
text list "Disconnect Code Descriptions Long": 0 'Connection terminated successfully.'; 28672 'No job processing active.'; 28673 'Start of job processing, connection being terminated.'; 28674 'Intermediate call (REQ irrelevant), connection being terminated.'; 32902 'The ID parameter is not in the permitted value range.'; 32931 'Attempt is being made to terminate a non-existent connection or the connection is already terminated.'; 32964 'Temporary communication error: New parameters are being assigned to the interface or the connection is currently being established.'; 65535 'In connect state.'

text list "Send Code Descriptions Long": 0 'Send job completed without error.'; 28672 'No job processing active.'; 28673 'Start of job execution, data is being sent. When processing this job, the operating system accesses the data in the DATA send area.'; 28674 'Job executing (REQ irrelevant). When processing this job, the operating system accesses the data in the DATA send area.'; 32901 'The LEN parameter is greater than the highest permitted value (65536). DATA and LEN parameters both have the value "0".'; 32902 'The ID parameter is outside the permitted address range (1..0xFFF).'; 32904 'The LEN parameter is greater than the area specified in DATA.'; 32929 'Communication error: The specified connection has not yet been established. The specified connection is being terminated. Transfer via thisconnection is not possible. The interface is being re-initialized.'; 32947 'The protocol variant (ConnectionType parameter in the connection description) is set to UDP. Use the instruction "TUSEND" with a UDP connection.'; 32963 'A block with this ID is already being processed in a different priority group. Internal lack of resources.'; 32964 'Temporary communication error: The connection cannot be established to the partner at this time. The interface is receiving new parameter settings or the connection is being established.'; 32965 'Connection terminated by the communication partner.'; 32966 'Network error. Communication partner cannot be reached.'; 32967 'Execution timeout'; 65535 'Function not yet called.'

text list "Status Lists": 0 ''; 1 ''; 2 ''; 3 ''

ScreenModuleEditorView "Connection_Status_Details" 790x405
   SymbolicIOField "header" at 0,0 size 790x50; TextOn '1'; TextOff '0'; TextList "Connection Details Header"
      Appearance <- "interface.header_animate"
      Visibility <- "interface.header_visible"
      ProcessValue <- "interface.header_selector"
   IOField "payload" at 0,55 size 790x295; FormatPattern ?????????????????????????????????????????????????????????????????????????????????????????????????????????????????????????????????????????????????????????????????????????????????????????????????????????????????????????????????????????????????????????????
      ProcessValue <- "interface.payload_text"
      Appearance <- "interface.payload_animate"
      Visibility <- "interface.payload_visible"
   Button "display_payload_button" at 0,355 size 790x50; TextOff 'DISPLAY PAYLOAD'
      Appearance <- "interface.display_payload_button_animate"
      ObjectEnable <- "interface.display_payload_button_enable"
      Visibility <- "interface.display_payload_button_visible"
      on Press: function_b14e0dd5("interface.display_payload_button_actuate", 0)
   SymbolicIOField "detailed_status" at 0,55 size 790x295; TextOff '0'; TextOn '1'; TextList "Status Lists"
      ProcessValue <- "interface.detailed_status_list_selector"
      Visibility <- "interface.detailed_status_visible"
      Appearance <- "interface.detailed_status_animate"
   Button "back_button" at 0,0 size 790x405; TextOff 'Text'
      ObjectEnable <- "interface.back_button_enable"
      Visibility <- "interface.back_button_visible"
      on Press: function_b14e0dd5("interface.back_button_actuate", 0)
*)

(* ===== HMI "HMI_RT_1" =====
system functions are stored by id; their names below are inferred from use

text list "Connection Details Header": 0 'NO STATE'; 1 'DISCONNECTION STATUS'; 2 'CONNECTION STATUS'; 3 'SEND STATUS'

text list "Connect Code Descriptions Long": 0 'Connection successfully established.'; 28672 'No job processing active'; 28673 'Start job execution, establish connection.'; 28674 'Connection is being established (REQ irrelevant).'; 32901 'Connection ID (ID parameter) is already being used by a configured connection.'; 32902 'The ID parameter is outside the valid range.'; 32903 'Maximum number of connections reached; no additional connection possible'; 32905 'The CONNECT parameter does not point to a data block.'; 32922 'The structure at the CONNECT parameter is not supported on an integrated interface or the length is invalid or an incorrect "InterfaceID" is specified in the connection description (SDT).'; 32923 'The element InterfaceId within the TCON_xxx structure does not reference a hardware identifier of a CPU or CM/CP interface or has the value "0".'; 32928 'Group error for error codes W#16#80A1 and W#16#80A2.'; 32929 'The specified connection or the port is already being used.'; 32930 'Local or remote port is being used by the system.'; 32931 'Attempt being made to re-establish an existing connection.'; 32932 'IP address of the remote endpoint of the connection is invalid, in other words, it matches the IP address of the local partner.'; 32933 'Connection ID is already in use.'; 32935 'Communication error: You executed "TDISCON" before "TCON" had completed.'; 32946 'The CONNECT parameter points to a data block that was generated with the attribute "Only store in load memory".'; 32948 'ISO-on-TCP violation: local_tsap_id_len >= B#16#02 local_tsap_id[1] = B#16#E0 local_tsap_id_len >= B#16#03 local_tsap_id[1] is ASCII chr local_tsap_id[1] is ASCII cha and local_tsap_id_len >= B#16#03'; 32949 'Only passive connection establishment is permitted for connection type 13 = UDP.'; 32950 'Parameter assignment error at the connection_type parameter of the SDT TCON_Param.'; 32951 'Error in one of the following parameters of the data block for connection description: block_length, local_tsap_id_len, rem_subnet_id_len, rem_staddr_len, rem_tsap_id_len, next_staddr_len. Note: If you call TCON in TCP for the passive end, local_tsap_id_len must have the value 2 and rem_tsap_id_len the value 0.'; 32952 'Connection description of the structure element ID and the block parameter ID are not identical.'; 32963 'All connection resources are in use.'; 32964 'Temporary communication error: Firewall Pending Parameterization Pending Disconnect'; 65535 'In disconnect state.'; 32966 'The connection partner could not be reached.'

text list "Disconnect Code Descriptions Long": 0 'Connection terminated successfully.'; 28672 'No job processing active.'; 28673 'Start of job processing, connection being terminated.'; 28674 'Intermediate call (REQ irrelevant), connection being terminated.'; 32902 'The ID parameter is not in the permitted value range.'; 32931 'Attempt is being made to terminate a non-existent connection or the connection is already terminated.'; 32964 'Temporary communication error: New parameters are being assigned to the interface or the connection is currently being established.'; 65535 'In connect state.'

text list "Send Code Descriptions Long": 0 'Send job completed without error.'; 28672 'No job processing active.'; 28673 'Start of job execution, data is being sent. When processing this job, the operating system accesses the data in the DATA send area.'; 28674 'Job executing (REQ irrelevant). When processing this job, the operating system accesses the data in the DATA send area.'; 32901 'The LEN parameter is greater than the highest permitted value (65536). DATA and LEN parameters both have the value "0".'; 32902 'The ID parameter is outside the permitted address range (1..0xFFF).'; 32904 'The LEN parameter is greater than the area specified in DATA.'; 32929 'Communication error: The specified connection has not yet been established. The specified connection is being terminated. Transfer via thisconnection is not possible. The interface is being re-initialized.'; 32947 'The protocol variant (ConnectionType parameter in the connection description) is set to UDP. Use the instruction "TUSEND" with a UDP connection.'; 32963 'A block with this ID is already being processed in a different priority group. Internal lack of resources.'; 32964 'Temporary communication error: The connection cannot be established to the partner at this time. The interface is receiving new parameter settings or the connection is being established.'; 32965 'Connection terminated by the communication partner.'; 32966 'Network error. Communication partner cannot be reached.'; 32967 'Execution timeout'; 65535 'Function not yet called.'

text list "Status Lists": 0 ''; 1 ''; 2 ''; 3 ''

ScreenModuleEditorView "Connection_Status_Details" 790x405
   SymbolicIOField "header" at 0,0 size 790x50; TextOn '1'; TextOff '0'; TextList "Connection Details Header"
      Appearance <- "interface.header_animate"
      Visibility <- "interface.header_visible"
      ProcessValue <- "interface.header_selector"
   IOField "payload" at 0,55 size 790x295; FormatPattern ?????????????????????????????????????????????????????????????????????????????????????????????????????????????????????????????????????????????????????????????????????????????????????????????????????????????????????????????????????????????????????????????
      Appearance <- "interface.payload_animate"
      ProcessValue <- "interface.payload_text"
      Visibility <- "interface.payload_visible"
   Button "display_payload_button" at 0,355 size 790x50; TextOff 'DISPLAY PAYLOAD'
      on Press: function_b14e0dd5("interface.display_payload_button_actuate", 0)
      Appearance <- "interface.display_payload_button_animate"
      ObjectEnable <- "interface.display_payload_button_enable"
      Visibility <- "interface.display_payload_button_visible"
   SymbolicIOField "detailed_status" at 0,55 size 790x295; TextOn '1'; TextOff '0'; TextList "Status Lists"
      Visibility <- "interface.detailed_status_visible"
      ProcessValue <- "interface.detailed_status_list_selector"
      Appearance <- "interface.detailed_status_animate"
   Button "back_button" at 0,0 size 790x405; TextOff 'Text'
      on Press: function_b14e0dd5("interface.back_button_actuate", 0)
      Visibility <- "interface.back_button_visible"
      ObjectEnable <- "interface.back_button_enable"
*)

(* ===== HMI "HMI_RT_1" =====
system functions are stored by id; their names below are inferred from use

text list "Connection Details Header": 0 'NO STATE'; 1 'DISCONNECTION STATUS'; 2 'CONNECTION STATUS'; 3 'SEND STATUS'

text list "Connect Code Descriptions Long": 0 'Connection successfully established.'; 28672 'No job processing active'; 28673 'Start job execution, establish connection.'; 28674 'Connection is being established (REQ irrelevant).'; 32901 'Connection ID (ID parameter) is already being used by a configured connection.'; 32902 'The ID parameter is outside the valid range.'; 32903 'Maximum number of connections reached; no additional connection possible'; 32905 'The CONNECT parameter does not point to a data block.'; 32922 'The structure at the CONNECT parameter is not supported on an integrated interface or the length is invalid or an incorrect "InterfaceID" is specified in the connection description (SDT).'; 32923 'The element InterfaceId within the TCON_xxx structure does not reference a hardware identifier of a CPU or CM/CP interface or has the value "0".'; 32928 'Group error for error codes W#16#80A1 and W#16#80A2.'; 32929 'The specified connection or the port is already being used.'; 32930 'Local or remote port is being used by the system.'; 32931 'Attempt being made to re-establish an existing connection.'; 32932 'IP address of the remote endpoint of the connection is invalid, in other words, it matches the IP address of the local partner.'; 32933 'Connection ID is already in use.'; 32935 'Communication error: You executed "TDISCON" before "TCON" had completed.'; 32946 'The CONNECT parameter points to a data block that was generated with the attribute "Only store in load memory".'; 32948 'ISO-on-TCP violation: local_tsap_id_len >= B#16#02 local_tsap_id[1] = B#16#E0 local_tsap_id_len >= B#16#03 local_tsap_id[1] is ASCII chr local_tsap_id[1] is ASCII cha and local_tsap_id_len >= B#16#03'; 32949 'Only passive connection establishment is permitted for connection type 13 = UDP.'; 32950 'Parameter assignment error at the connection_type parameter of the SDT TCON_Param.'; 32951 'Error in one of the following parameters of the data block for connection description: block_length, local_tsap_id_len, rem_subnet_id_len, rem_staddr_len, rem_tsap_id_len, next_staddr_len. Note: If you call TCON in TCP for the passive end, local_tsap_id_len must have the value 2 and rem_tsap_id_len the value 0.'; 32952 'Connection description of the structure element ID and the block parameter ID are not identical.'; 32963 'All connection resources are in use.'; 32964 'Temporary communication error: Firewall Pending Parameterization Pending Disconnect'; 65535 'In disconnect state.'; 32966 'The connection partner could not be reached.'

text list "Disconnect Code Descriptions Long": 0 'Connection terminated successfully.'; 28672 'No job processing active.'; 28673 'Start of job processing, connection being terminated.'; 28674 'Intermediate call (REQ irrelevant), connection being terminated.'; 32902 'The ID parameter is not in the permitted value range.'; 32931 'Attempt is being made to terminate a non-existent connection or the connection is already terminated.'; 32964 'Temporary communication error: New parameters are being assigned to the interface or the connection is currently being established.'; 65535 'In connect state.'

text list "Send Code Descriptions Long": 0 'Send job completed without error.'; 28672 'No job processing active.'; 28673 'Start of job execution, data is being sent. When processing this job, the operating system accesses the data in the DATA send area.'; 28674 'Job executing (REQ irrelevant). When processing this job, the operating system accesses the data in the DATA send area.'; 32901 'The LEN parameter is greater than the highest permitted value (65536). DATA and LEN parameters both have the value "0".'; 32902 'The ID parameter is outside the permitted address range (1..0xFFF).'; 32904 'The LEN parameter is greater than the area specified in DATA.'; 32929 'Communication error: The specified connection has not yet been established. The specified connection is being terminated. Transfer via thisconnection is not possible. The interface is being re-initialized.'; 32947 'The protocol variant (ConnectionType parameter in the connection description) is set to UDP. Use the instruction "TUSEND" with a UDP connection.'; 32963 'A block with this ID is already being processed in a different priority group. Internal lack of resources.'; 32964 'Temporary communication error: The connection cannot be established to the partner at this time. The interface is receiving new parameter settings or the connection is being established.'; 32965 'Connection terminated by the communication partner.'; 32966 'Network error. Communication partner cannot be reached.'; 32967 'Execution timeout'; 65535 'Function not yet called.'

text list "Status Lists": 0 ''; 1 ''; 2 ''; 3 ''

ScreenModuleEditorView "Connection_Status_Details" 790x405
   SymbolicIOField "header" at 0,0 size 790x50; TextOn '1'; TextOff '0'; TextList "Connection Details Header"
      Appearance <- "interface.header_animate"
      Visibility <- "interface.header_visible"
      ProcessValue <- "interface.header_selector"
   IOField "payload" at 0,55 size 790x295; FormatPattern ?????????????????????????????????????????????????????????????????????????????????????????????????????????????????????????????????????????????????????????????????????????????????????????????????????????????????????????????????????????????????????????????
      Appearance <- "interface.payload_animate"
      ProcessValue <- "interface.payload_text"
      Visibility <- "interface.payload_visible"
   Button "display_payload_button" at 0,355 size 790x50; TextOff 'DISPLAY PAYLOAD'
      on Press: function_b14e0dd5("interface.display_payload_button_actuate", 0)
      Appearance <- "interface.display_payload_button_animate"
      ObjectEnable <- "interface.display_payload_button_enable"
      Visibility <- "interface.display_payload_button_visible"
   SymbolicIOField "detailed_status" at 0,55 size 790x295; TextOn '1'; TextOff '0'; TextList "Status Lists"
      Visibility <- "interface.detailed_status_visible"
      ProcessValue <- "interface.detailed_status_list_selector"
      Appearance <- "interface.detailed_status_animate"
   Button "back_button" at 0,0 size 790x405; TextOff 'Text'
      on Press: function_b14e0dd5("interface.back_button_actuate", 0)
      Visibility <- "interface.back_button_visible"
      ObjectEnable <- "interface.back_button_enable"
*)

(* ===== HMI "HMI_RT_1" =====
system functions are stored by id; their names below are inferred from use

text list "Send Code Descriptions Short": 0 'SEND SUCCESSFUL'; 28672 'NO JOB'; 28673 'DATA ACCESSED DURING JOB'; 28674 'JOB PROCESSING'; 32901 'MAX LENGTH EXCEEDED'; 32902 'INVALID ID OUT OF RANGE'; 32904 'LENGTH EXCEEDS DATA RANGE'; 32929 'NO CONNECTION'; 32947 'UDP CONNECTION'; 32963 'CONNECTION BUSY'; 32964 'REQUEST DURING PARAM ASSIGNMENT'; 32965 'PARTNER TERMINATED CONNECTION'; 32966 'PARTNER UNAVAILABLE'; 32967 'TIMEOUT'; 65535 'NOT CALLED'

text list "Connect Code Descriptions Short": 0 'CONNECTION SUCCESSFUL'; 28672 'NO JOB'; 28673 'START JOB'; 28674 'PROCESSING JOB'; 32901 'ID INVALID: ALREADY IN USE'; 32902 'ID INVALID: OUT OF RANGE'; 32903 'MAX CONNECTIONS REACHED'; 32905 'NO CONNECTION DATA STORED'; 32922 'INVALID CONNECTION DATA'; 32923 'NO CONNECTION HARDWARE'; 32928 'GROUP ERROR'; 32929 'LOCAL PORT IN USE'; 32930 'REMOTE PORT IN USE'; 32931 'CONNECTION ALREADY ESTABLISHED'; 32932 'INVALID IP ADDRESS'; 32933 'DUPLICATE CONNECTION ID'; 32935 'DICONNECT REQUEST WHILE CONNECTING'; 32946 'CONNECT DATA IN LOAD MEMORY'; 32948 'ISO ON TCP VIOLATION'; 32949 'NON PASSIVE UDP CONNECTION REQUEST'; 32950 'INVALID CONNECTION TYPE'; 32951 'CONNECTION PARAMETER ERROR'; 32952 'DATA/PARAMETER MISMATCH'; 32963 'MAX CONNECTIONS EXCEEDED'; 32964 'FIREWALL'; 65535 'STATE: DISCONNECT'; 32966 'PARTNER UNAVAILABLE'

text list "Disconnect Code Descriptions Short": 0 'DISCONNECTION SUCCESSFUL'; 28672 'NO JOB'; 28673 'JOB STARTED'; 28674 'REQUEST DURING EXECUTION'; 32902 'ID INVALID: OUT OF RANGE'; 32931 'CONNECTION ALREADY TERMINATED'; 32964 'REQUEST DURING PARAM ASSIGNMENT'; 65535 'STATE: CONNECT'

text list "Text List Select": 0 ''; 1 ''; 2 ''; 3 ''

ScreenModuleEditorView "Connection_Status_Element" 392x110
   TextField "operation_label" at 0,0 size 110x110; Text 'S'
      Visibility <- "interface.operation_label_visible"
      Appearance <- "interface.operation_label_animate"
   TextField "done_status_indicator" at 110,0 size 94x27; Text 'DONE'
      Visibility <- "interface.done_status_indicator_visible"
      Appearance <- "interface.done_status_indicator_animate"
   TextField "busy_status_indicator" at 204,0 size 94x27; Text 'BUSY'
      Visibility <- "interface.busy_status_indicator_visible"
      Appearance <- "interface.busy_status_indicator_animate"
   TextField "error_status_indicator" at 298,0 size 94x27; Text 'ERROR'
      Visibility <- "interface.error_status_indicator_visible"
      Appearance <- "interface.error_status_indicator_animate"
   TextField "status_code_label" at 110,27 size 82x28; Text 'CODE:'
      Visibility <- "interface.status_code_label_visible"
      Appearance <- "interface.status_code_label_animate"
   IOField "status_code" at 192,27 size 200x28; FormatPattern ??????
      Appearance <- "interface.status_code_value_animate"
      Visibility <- "interface.status_code_value_visible"
      ProcessValue <- "interface.status_code_value"
   SymbolicIOField "status_description" at 110,55 size 282x55; TextOn '1'; TextOff '0'; TextList "Text List Select"
      Appearance <- "interface.status_code_description_animate"
      ProcessValue <- "operation_list_selector"
      Visibility <- "interface.status_code_description_visible"
   Button "operation_left" at 0,0 size 110x110; TextOff 'Text'
      on Press: function_b14e0dd5("interface.operation_button_actuate", 0)
      Visibility <- "interface.operation_button_visible"
      ObjectEnable <- "interface.operation_button_enable"
   Button "operation_top" at 110,0 size 282x55; TextOff 'Text'
      on Press: function_b14e0dd5("interface.operation_button_actuate", 0)
      Visibility <- "interface.operation_button_visible"
      ObjectEnable <- "interface.operation_button_enable"
   Button "show_status" at 110,55 size 282x55; TextOff 'Text'
      on Press: function_b14e0dd5("interface.show_status_code_description_button_actuate", 0)
      Visibility <- "interface.show_status_code_description_button_visible"
      ObjectEnable <- "interface.show_status_code_description_button_enable"
*)

(* ===== HMI "HMI_RT_1" =====
system functions are stored by id; their names below are inferred from use

text list "Send Code Descriptions Short": 0 'SEND SUCCESSFUL'; 28672 'NO JOB'; 28673 'DATA ACCESSED DURING JOB'; 28674 'JOB PROCESSING'; 32901 'MAX LENGTH EXCEEDED'; 32902 'INVALID ID OUT OF RANGE'; 32904 'LENGTH EXCEEDS DATA RANGE'; 32929 'NO CONNECTION'; 32947 'UDP CONNECTION'; 32963 'CONNECTION BUSY'; 32964 'REQUEST DURING PARAM ASSIGNMENT'; 32965 'PARTNER TERMINATED CONNECTION'; 32966 'PARTNER UNAVAILABLE'; 32967 'TIMEOUT'; 65535 'NOT CALLED'; -1 'NO STATE'

text list "Connect Code Descriptions Short": 0 'CONNECTION SUCCESSFUL'; 28672 'NO JOB'; 28673 'START JOB'; 28674 'PROCESSING JOB'; 32901 'ID INVALID: ALREADY IN USE'; 32902 'ID INVALID: OUT OF RANGE'; 32903 'MAX CONNECTIONS REACHED'; 32905 'NO CONNECTION DATA STORED'; 32922 'INVALID CONNECTION DATA'; 32923 'NO CONNECTION HARDWARE'; 32928 'GROUP ERROR'; 32929 'LOCAL PORT IN USE'; 32930 'REMOTE PORT IN USE'; 32931 'CONNECTION ALREADY ESTABLISHED'; 32932 'INVALID IP ADDRESS'; 32933 'DUPLICATE CONNECTION ID'; 32935 'DICONNECT REQUEST WHILE CONNECTING'; 32946 'CONNECT DATA IN LOAD MEMORY'; 32948 'ISO ON TCP VIOLATION'; 32949 'NON PASSIVE UDP CONNECTION REQUEST'; 32950 'INVALID CONNECTION TYPE'; 32951 'CONNECTION PARAMETER ERROR'; 32952 'DATA/PARAMETER MISMATCH'; 32963 'MAX CONNECTIONS EXCEEDED'; 32964 'FIREWALL'; 65535 'STATE: DISCONNECT'; 32966 'PARTNER UNAVAILABLE'; -1 'NO STATE'

text list "Disconnect Code Descriptions Short": 0 'DISCONNECTION SUCCESSFUL'; 28672 'NO JOB'; 28673 'JOB STARTED'; 28674 'REQUEST DURING EXECUTION'; 32902 'ID INVALID: OUT OF RANGE'; 32931 'CONNECTION ALREADY TERMINATED'; 32964 'REQUEST DURING PARAM ASSIGNMENT'; 65535 'STATE: CONNECT'; -1 'NO STATE'

text list "Text List Select": 0 ''; 1 ''; 2 ''; 3 ''

ScreenModuleEditorView "Connection_Status_Element" 392x110
   TextField "operation_label" at 0,0 size 110x110; Text 'S'
      Visibility <- "interface.operation_label_visible"
      Appearance <- "interface.operation_label_animate"
   TextField "done_status_indicator" at 110,0 size 94x27; Text 'DONE'
      Visibility <- "interface.done_status_indicator_visible"
      Appearance <- "interface.done_status_indicator_animate"
   TextField "busy_status_indicator" at 204,0 size 94x27; Text 'BUSY'
      Visibility <- "interface.busy_status_indicator_visible"
      Appearance <- "interface.busy_status_indicator_animate"
   TextField "error_status_indicator" at 298,0 size 94x27; Text 'ERROR'
      Visibility <- "interface.error_status_indicator_visible"
      Appearance <- "interface.error_status_indicator_animate"
   TextField "status_code_label" at 110,27 size 82x28; Text 'CODE:'
      Visibility <- "interface.status_code_label_visible"
      Appearance <- "interface.status_code_label_animate"
   IOField "status_code" at 192,27 size 200x28; FormatPattern ??????
      Appearance <- "interface.status_code_value_animate"
      Visibility <- "interface.status_code_value_visible"
      ProcessValue <- "interface.status_code_value"
   SymbolicIOField "status_description" at 110,55 size 282x55; TextOn '1'; TextOff '0'; TextList "Text List Select"
      Appearance <- "interface.status_code_description_animate"
      ProcessValue <- "operation_list_selector"
      Visibility <- "interface.status_code_description_visible"
   Button "operation_left" at 0,0 size 110x110; TextOff 'Text'
      on Press: function_b14e0dd5("interface.operation_button_actuate", 0)
      Visibility <- "interface.operation_button_visible"
      ObjectEnable <- "interface.operation_button_enable"
   Button "operation_top" at 110,0 size 282x55; TextOff 'Text'
      on Press: function_b14e0dd5("interface.operation_button_actuate", 0)
      Visibility <- "interface.operation_button_visible"
      ObjectEnable <- "interface.operation_button_enable"
   Button "show_status" at 110,55 size 282x55; TextOff 'Text'
      on Press: function_b14e0dd5("interface.show_status_code_description_button_actuate", 0)
      Visibility <- "interface.show_status_code_description_button_visible"
      ObjectEnable <- "interface.show_status_code_description_button_enable"
*)

(* ===== HMI "HMI_RT_1" =====
system functions are stored by id; their names below are inferred from use

text list "Send Code Descriptions Short": 0 'SEND SUCCESSFUL'; 28672 'NO JOB'; 28673 'DATA ACCESSED DURING JOB'; 28674 'JOB PROCESSING'; 32901 'MAX LENGTH EXCEEDED'; 32902 'INVALID ID OUT OF RANGE'; 32904 'LENGTH EXCEEDS DATA RANGE'; 32929 'NO CONNECTION'; 32947 'UDP CONNECTION'; 32963 'CONNECTION BUSY'; 32964 'REQUEST DURING PARAM ASSIGNMENT'; 32965 'PARTNER TERMINATED CONNECTION'; 32966 'PARTNER UNAVAILABLE'; 32967 'TIMEOUT'; 65535 'NOT CALLED'; -1 'NO STATE'

text list "Connect Code Descriptions Short": 0 'CONNECTION SUCCESSFUL'; 28672 'NO JOB'; 28673 'START JOB'; 28674 'PROCESSING JOB'; 32901 'ID INVALID: ALREADY IN USE'; 32902 'ID INVALID: OUT OF RANGE'; 32903 'MAX CONNECTIONS REACHED'; 32905 'NO CONNECTION DATA STORED'; 32922 'INVALID CONNECTION DATA'; 32923 'NO CONNECTION HARDWARE'; 32928 'GROUP ERROR'; 32929 'LOCAL PORT IN USE'; 32930 'REMOTE PORT IN USE'; 32931 'CONNECTION ALREADY ESTABLISHED'; 32932 'INVALID IP ADDRESS'; 32933 'DUPLICATE CONNECTION ID'; 32935 'DICONNECT REQUEST WHILE CONNECTING'; 32946 'CONNECT DATA IN LOAD MEMORY'; 32948 'ISO ON TCP VIOLATION'; 32949 'NON PASSIVE UDP CONNECTION REQUEST'; 32950 'INVALID CONNECTION TYPE'; 32951 'CONNECTION PARAMETER ERROR'; 32952 'DATA/PARAMETER MISMATCH'; 32963 'MAX CONNECTIONS EXCEEDED'; 32964 'FIREWALL'; 65535 'STATE: DISCONNECT'; 32966 'PARTNER UNAVAILABLE'; -1 'NO STATE'

text list "Disconnect Code Descriptions Short": 0 'DISCONNECTION SUCCESSFUL'; 28672 'NO JOB'; 28673 'JOB STARTED'; 28674 'REQUEST DURING EXECUTION'; 32902 'ID INVALID: OUT OF RANGE'; 32931 'CONNECTION ALREADY TERMINATED'; 32964 'REQUEST DURING PARAM ASSIGNMENT'; 65535 'STATE: CONNECT'; -1 'NO STATE'

text list "Text List Select": 0 ''; 1 ''; 2 ''; 3 ''

ScreenModuleEditorView "Connection_Status_Element" 392x110
   TextField "operation_label" at 0,0 size 110x110; Text 'S'
      Visibility <- "interface.operation_label_visible"
      Appearance <- "interface.operation_label_animate"
   TextField "done_status_indicator" at 110,0 size 94x27; Text 'DONE'
      Visibility <- "interface.done_status_indicator_visible"
      Appearance <- "interface.done_status_indicator_animate"
   TextField "busy_status_indicator" at 204,0 size 94x27; Text 'BUSY'
      Visibility <- "interface.busy_status_indicator_visible"
      Appearance <- "interface.busy_status_indicator_animate"
   TextField "error_status_indicator" at 298,0 size 94x27; Text 'ERROR'
      Visibility <- "interface.error_status_indicator_visible"
      Appearance <- "interface.error_status_indicator_animate"
   TextField "status_code_label" at 110,27 size 82x28; Text 'CODE:'
      Visibility <- "interface.status_code_label_visible"
      Appearance <- "interface.status_code_label_animate"
   IOField "status_code" at 192,27 size 200x28; FormatPattern ??????
      Appearance <- "interface.status_code_value_animate"
      Visibility <- "interface.status_code_value_visible"
      ProcessValue <- "interface.status_code_value"
   SymbolicIOField "status_description" at 110,55 size 282x55; TextOn '1'; TextOff '0'; TextList "Text List Select"
      Appearance <- "interface.status_code_description_animate"
      ProcessValue <- "operation_list_selector"
      Visibility <- "interface.status_code_description_visible"
   Button "operation_left" at 0,0 size 110x110; TextOff 'Text'
      on Press: function_b14e0dd5("interface.operation_button_actuate", 0)
      Visibility <- "interface.operation_button_visible"
      ObjectEnable <- "interface.operation_button_enable"
   Button "operation_top" at 110,0 size 282x55; TextOff 'Text'
      on Press: function_b14e0dd5("interface.operation_button_actuate", 0)
      Visibility <- "interface.operation_button_visible"
      ObjectEnable <- "interface.operation_button_enable"
   Button "show_status" at 110,55 size 282x55; TextOff 'Text'
      on Press: function_b14e0dd5("interface.show_status_code_description_button_actuate", 0)
      Visibility <- "interface.show_status_code_description_button_visible"
      ObjectEnable <- "interface.show_status_code_description_button_enable"
*)

(* ===== HMI "HMI_RT_1" =====
system functions are stored by id; their names below are inferred from use

ScreenModuleEditorView "Connection_Parameters_Control" 600x270
   TextField "id_label" at 0,55 size 300x50; Text 'ID'
      Appearance <- "interface.id_label_animate"
      Visibility <- "interface.id_label_visible"
   IOField "id_entry" at 300,55 size 300x50; FormatPattern ??????
      Appearance <- "interface.id_entry_animate"
      Visibility <- "interface.id_entry_visible"
      ObjectEnable <- "interface.id_entry_enable"
      ProcessValue <- "interface.id_entry_value"
   Button "back" at 0,220 size 600x50; TextOff 'BACK'
      Appearance <- "interface.back_animate"
      Visibility <- "interface.back_visible"
      ObjectEnable <- "interface.back_enable"
      on Press: function_b14e0dd5("interface.back_actuate", 0)
   TextField "ip_address_label" at 0,110 size 300x50; Text 'IP ADDRESS'
      Appearance <- "interface.ip_address_label_animate"
      Visibility <- "interface.ip_address_label_visible"
   IOField "ip_address_entry" at 300,110 size 300x50; FormatPattern ???????????????
      Appearance <- "interface.ip_address_entry_animate"
      Visibility <- "interface.ip_address_entry_visible"
      ObjectEnable <- "interface.ip_address_entry_enable"
      ProcessValue <- "interface.ip_address_entry_value"
   TextField "port_label" at 0,165 size 300x50; Text 'PORT'
      Appearance <- "interface.port_label_animate"
      Visibility <- "interface.port_label_visible"
   IOField "port_entry" at 300,165 size 300x50; FormatPattern ??????
      Appearance <- "interface.port_entry_animate"
      Visibility <- "interface.port_entry_visible"
      ObjectEnable <- "interface.port_entry_enable"
      ProcessValue <- "interface.port_entry_value"
   IOField "I/O field_1" at 0,0 size 600x50; FormatPattern ?????????????????????????
      Appearance <- "interface.header_animate"
      Visibility <- "interface.header_visible"
*)

(* ===== HMI "HMI_RT_1" =====
system functions are stored by id; their names below are inferred from use

ScreenModuleEditorView "Connection_Status_Header" 392x55
   Button "header" at 0,0 size 392x55; TextOff 'PARTNER CONNECTION CONTROLS'
      Visibility <- "interface.visible"
      Appearance <- "interface.animate"
      on Press: function_b14e0dd5("interface.actuate", 0)
      ObjectEnable <- "interface.enable"
*)

(* ===== HMI "HMI_RT_1" =====
system functions are stored by id; their names below are inferred from use

ScreenModuleEditorView "Connection_Parameters_Control" 600x270
   TextField "id_label" at 0,55 size 300x50; Text 'ID'
      Visibility <- "interface.id_label_visible"
      Appearance <- "interface.id_label_animate"
   IOField "id_entry" at 300,55 size 300x50; FormatPattern ??????
      Appearance <- "interface.id_entry_animate"
      Visibility <- "interface.id_entry_visible"
      ProcessValue <- "interface.id_entry_value"
      ObjectEnable <- "interface.id_entry_enable"
   Button "back" at 0,220 size 600x50; TextOff 'BACK'
      on Press: function_b14e0dd5("interface.back_actuate", 0)
      Appearance <- "interface.back_animate"
      Visibility <- "interface.back_visible"
      ObjectEnable <- "interface.back_enable"
   TextField "ip_address_label" at 0,110 size 300x50; Text 'IP ADDRESS'
      Visibility <- "interface.ip_address_label_visible"
      Appearance <- "interface.ip_address_label_animate"
   IOField "ip_address_entry" at 300,110 size 300x50; FormatPattern ???????????????
      Appearance <- "interface.ip_address_entry_animate"
      Visibility <- "interface.ip_address_entry_visible"
      ProcessValue <- "interface.ip_address_entry_value"
      ObjectEnable <- "interface.ip_address_entry_enable"
   TextField "port_label" at 0,165 size 300x50; Text 'PORT'
      Visibility <- "interface.port_label_visible"
      Appearance <- "interface.port_label_animate"
   IOField "port_entry" at 300,165 size 300x50; FormatPattern ??????
      Appearance <- "interface.port_entry_animate"
      Visibility <- "interface.port_entry_visible"
      ProcessValue <- "interface.port_entry_value"
      ObjectEnable <- "interface.port_entry_enable"
   IOField "header" at 0,0 size 600x50; FormatPattern ?????????????????????????
      Visibility <- "interface.header_visible"
      Appearance <- "interface.header_animate"
      ProcessValue <- "interface.header_value"
*)

(* ===== HMI "HMI_RT_1" =====
system functions are stored by id; their names below are inferred from use

ScreenModuleEditorView "Connection_Status_Header" 392x55
   Button "header" at 0,0 size 392x55; TextOff 'PARTNER CONNECTION CONTROLS'
      on Press: function_b14e0dd5("interface.actuate", 0)
      Appearance <- "interface.animate"
      Visibility <- "interface.visible"
      ObjectEnable <- "interface.enable"
*)

(* ===== HMI "HMI_RT_1" =====
system functions are stored by id; their names below are inferred from use

ScreenModuleEditorView "Connection_Status_Header" 392x55
   Button "header" at 0,0 size 392x55; TextOff 'PARTNER CONNECTION CONTROLS'
      on Press: function_b14e0dd5("interface.actuate", 0)
      Appearance <- "interface.animate"
      Visibility <- "interface.visible"
      ObjectEnable <- "interface.enable"
*)

(* ===== HMI "HMI_RT_1" =====
system functions are stored by id; their names below are inferred from use

ScreenModuleEditorView "Connection_Parameters_Control" 600x270
   TextField "id_label" at 0,55 size 300x50; Text 'ID'
      Visibility <- "interface.id_label_visible"
      Appearance <- "interface.id_label_animate"
   IOField "id_entry" at 300,55 size 300x50; FormatPattern ??????
      Appearance <- "interface.id_entry_animate"
      Visibility <- "interface.id_entry_visible"
      ObjectEnable <- "interface.id_entry_enable"
      ProcessValue <- "interface.id_entry_value"
      on OnFinishInput: SetBit("interface.id_entry_input_finished")
   Button "back" at 0,220 size 600x50; TextOff 'BACK'
      on Press: function_b14e0dd5("interface.back_actuate", 0)
      Appearance <- "interface.back_animate"
      Visibility <- "interface.back_visible"
      ObjectEnable <- "interface.back_enable"
   TextField "ip_address_label" at 0,110 size 300x50; Text 'IP ADDRESS'
      Visibility <- "interface.ip_address_label_visible"
      Appearance <- "interface.ip_address_label_animate"
   IOField "ip_address_entry" at 300,110 size 300x50; FormatPattern ???????????????
      Appearance <- "interface.ip_address_entry_animate"
      Visibility <- "interface.ip_address_entry_visible"
      ObjectEnable <- "interface.ip_address_entry_enable"
      ProcessValue <- "interface.ip_address_entry_value"
      on OnFinishInput: SetBit("interface.ip_address_entry_input_finished")
   TextField "port_label" at 0,165 size 300x50; Text 'PORT'
      Visibility <- "interface.port_label_visible"
      Appearance <- "interface.port_label_animate"
   IOField "port_entry" at 300,165 size 300x50; FormatPattern ??????
      Appearance <- "interface.port_entry_animate"
      Visibility <- "interface.port_entry_visible"
      ObjectEnable <- "interface.port_entry_enable"
      ProcessValue <- "interface.port_entry_value"
      on OnFinishInput: SetBit("interface.port_entry_input_finished")
   IOField "header" at 0,0 size 600x50; FormatPattern ?????????????????????????
      Appearance <- "interface.header_animate"
      Visibility <- "interface.header_visible"
      ProcessValue <- "interface.header_value"
*)

(* ===== HMI "HMI_RT_1" =====
system functions are stored by id; their names below are inferred from use

ScreenModuleEditorView "Connection_Parameters_Control" 600x270
   TextField "id_label" at 0,55 size 300x50; Text 'ID'
      Visibility <- "interface.id_label_visible"
      Appearance <- "interface.id_label_animate"
   IOField "id_entry" at 300,55 size 300x50; FormatPattern ??????
      on OnFinishInput: SetBit("interface.id_entry_input_finished")
      Appearance <- "interface.id_entry_animate"
      Visibility <- "interface.id_entry_visible"
      ProcessValue <- "interface.id_entry_value"
      ObjectEnable <- "interface.id_entry_enable"
      on Activate: SetBit("interface.id_entry_active")
      on Deactivate: ResetBit("interface.id_entry_active")
   Button "back" at 0,220 size 600x50; TextOff 'BACK'
      on Press: function_b14e0dd5("interface.back_actuate", 0)
      Appearance <- "interface.back_animate"
      Visibility <- "interface.back_visible"
      ObjectEnable <- "interface.back_enable"
   TextField "ip_address_label" at 0,110 size 300x50; Text 'IP ADDRESS'
      Visibility <- "interface.ip_address_label_visible"
      Appearance <- "interface.ip_address_label_animate"
   IOField "ip_address_entry" at 300,110 size 300x50; FormatPattern ???????????????
      on OnFinishInput: SetBit("interface.ip_address_entry_input_finished")
      Appearance <- "interface.ip_address_entry_animate"
      Visibility <- "interface.ip_address_entry_visible"
      ProcessValue <- "interface.ip_address_entry_value"
      ObjectEnable <- "interface.ip_address_entry_enable"
      on Activate: SetBit("interface.ip_address_entry_active")
      on Deactivate: ResetBit("interface.ip_address_entry_active")
   TextField "port_label" at 0,165 size 300x50; Text 'PORT'
      Visibility <- "interface.port_label_visible"
      Appearance <- "interface.port_label_animate"
   IOField "port_entry" at 300,165 size 300x50; FormatPattern ??????
      on OnFinishInput: SetBit("interface.port_entry_input_finished")
      Appearance <- "interface.port_entry_animate"
      Visibility <- "interface.port_entry_visible"
      ProcessValue <- "interface.port_entry_value"
      ObjectEnable <- "interface.port_entry_enable"
      on Activate: SetBit("interface.port_entry_active")
      on Deactivate: ResetBit("interface.port_entry_active")
   IOField "header" at 0,0 size 600x50; FormatPattern ?????????????????????????
      Appearance <- "interface.header_animate"
      Visibility <- "interface.header_visible"
      ProcessValue <- "interface.header_value"
*)

(* ===== HMI "HMI_RT_1" =====
system functions are stored by id; their names below are inferred from use

text list "Send Code Descriptions Short": 0 'SEND SUCCESSFUL'; 28672 'NO JOB'; 28673 'DATA ACCESSED DURING JOB'; 28674 'JOB PROCESSING'; 32901 'MAX LENGTH EXCEEDED'; 32902 'INVALID ID OUT OF RANGE'; 32904 'LENGTH EXCEEDS DATA RANGE'; 32929 'NO CONNECTION'; 32947 'UDP CONNECTION'; 32963 'CONNECTION BUSY'; 32964 'REQUEST DURING PARAM ASSIGNMENT'; 32965 'PARTNER TERMINATED CONNECTION'; 32966 'PARTNER UNAVAILABLE'; 32967 'TIMEOUT'; 65535 'NOT CALLED'; -1 'NO STATE'

text list "Connect Code Descriptions Short": 0 'CONNECTION SUCCESSFUL'; 28672 'NO JOB'; 28673 'START JOB'; 28674 'PROCESSING JOB'; 32901 'ID INVALID: ALREADY IN USE'; 32902 'ID INVALID: OUT OF RANGE'; 32903 'MAX CONNECTIONS REACHED'; 32905 'NO CONNECTION DATA STORED'; 32922 'INVALID CONNECTION DATA'; 32923 'NO CONNECTION HARDWARE'; 32928 'GROUP ERROR'; 32929 'LOCAL PORT IN USE'; 32930 'REMOTE PORT IN USE'; 32931 'CONNECTION ALREADY ESTABLISHED'; 32932 'INVALID IP ADDRESS'; 32933 'DUPLICATE CONNECTION ID'; 32935 'DICONNECT REQUEST WHILE CONNECTING'; 32946 'CONNECT DATA IN LOAD MEMORY'; 32948 'ISO ON TCP VIOLATION'; 32949 'NON PASSIVE UDP CONNECTION REQUEST'; 32950 'INVALID CONNECTION TYPE'; 32951 'CONNECTION PARAMETER ERROR'; 32952 'DATA/PARAMETER MISMATCH'; 32963 'MAX CONNECTIONS EXCEEDED'; 32964 'FIREWALL'; 65535 'STATE: DISCONNECT'; 32966 'PARTNER UNAVAILABLE'; -1 'NO STATE'; 32965 'CONNECTION REFUSED'

text list "Disconnect Code Descriptions Short": 0 'DISCONNECTION SUCCESSFUL'; 28672 'NO JOB'; 28673 'JOB STARTED'; 28674 'REQUEST DURING EXECUTION'; 32902 'ID INVALID: OUT OF RANGE'; 32931 'CONNECTION ALREADY TERMINATED'; 32964 'REQUEST DURING PARAM ASSIGNMENT'; 65535 'STATE: CONNECT'; -1 'NO STATE'

text list "Text List Select": 0 ''; 1 ''; 2 ''; 3 ''

ScreenModuleEditorView "Connection_Status_Element" 392x110
   TextField "operation_label" at 0,0 size 110x110; Text 'S'
      Visibility <- "interface.operation_label_visible"
      Appearance <- "interface.operation_label_animate"
   TextField "done_status_indicator" at 110,0 size 94x27; Text 'DONE'
      Visibility <- "interface.done_status_indicator_visible"
      Appearance <- "interface.done_status_indicator_animate"
   TextField "busy_status_indicator" at 204,0 size 94x27; Text 'BUSY'
      Visibility <- "interface.busy_status_indicator_visible"
      Appearance <- "interface.busy_status_indicator_animate"
   TextField "error_status_indicator" at 298,0 size 94x27; Text 'ERROR'
      Visibility <- "interface.error_status_indicator_visible"
      Appearance <- "interface.error_status_indicator_animate"
   TextField "status_code_label" at 110,27 size 82x28; Text 'CODE:'
      Visibility <- "interface.status_code_label_visible"
      Appearance <- "interface.status_code_label_animate"
   IOField "status_code" at 192,27 size 200x28; FormatPattern ??????
      Appearance <- "interface.status_code_value_animate"
      Visibility <- "interface.status_code_value_visible"
      ProcessValue <- "interface.status_code_value"
   SymbolicIOField "status_description" at 110,55 size 282x55; TextOn '1'; TextOff '0'; TextList "Text List Select"
      Appearance <- "interface.status_code_description_animate"
      ProcessValue <- "operation_list_selector"
      Visibility <- "interface.status_code_description_visible"
   Button "operation_left" at 0,0 size 110x110; TextOff 'Text'
      on Press: function_b14e0dd5("interface.operation_button_actuate", 0)
      Visibility <- "interface.operation_button_visible"
      ObjectEnable <- "interface.operation_button_enable"
   Button "operation_top" at 110,0 size 282x55; TextOff 'Text'
      on Press: function_b14e0dd5("interface.operation_button_actuate", 0)
      Visibility <- "interface.operation_button_visible"
      ObjectEnable <- "interface.operation_button_enable"
   Button "show_status" at 110,55 size 282x55; TextOff 'Text'
      on Press: function_b14e0dd5("interface.show_status_code_description_button_actuate", 0)
      Visibility <- "interface.show_status_code_description_button_visible"
      ObjectEnable <- "interface.show_status_code_description_button_enable"
*)

(* ===== HMI "HMI_RT_1" =====
system functions are stored by id; their names below are inferred from use

text list "Send Code Descriptions Short": 0 'SEND SUCCESSFUL'; 28672 'NO JOB'; 28673 'DATA ACCESSED DURING JOB'; 28674 'JOB PROCESSING'; 32901 'MAX LENGTH EXCEEDED'; 32902 'INVALID ID OUT OF RANGE'; 32904 'LENGTH EXCEEDS DATA RANGE'; 32929 'NO CONNECTION'; 32947 'UDP CONNECTION'; 32963 'CONNECTION BUSY'; 32964 'REQUEST DURING PARAM ASSIGNMENT'; 32965 'PARTNER TERMINATED CONNECTION'; 32966 'PARTNER UNAVAILABLE'; 32967 'TIMEOUT'; 65535 'NOT CALLED'; -1 'NO STATE'

text list "Connect Code Descriptions Short": 0 'CONNECTION SUCCESSFUL'; 28672 'NO JOB'; 28673 'START JOB'; 28674 'PROCESSING JOB'; 32901 'ID INVALID: ALREADY IN USE'; 32902 'ID INVALID: OUT OF RANGE'; 32903 'MAX CONNECTIONS REACHED'; 32905 'NO CONNECTION DATA STORED'; 32922 'INVALID CONNECTION DATA'; 32923 'NO CONNECTION HARDWARE'; 32928 'GROUP ERROR'; 32929 'LOCAL PORT IN USE'; 32930 'REMOTE PORT IN USE'; 32931 'CONNECTION ALREADY ESTABLISHED'; 32932 'INVALID IP ADDRESS'; 32933 'DUPLICATE CONNECTION ID'; 32935 'DICONNECT REQUEST WHILE CONNECTING'; 32946 'CONNECT DATA IN LOAD MEMORY'; 32948 'ISO ON TCP VIOLATION'; 32949 'NON PASSIVE UDP CONNECTION REQUEST'; 32950 'INVALID CONNECTION TYPE'; 32951 'CONNECTION PARAMETER ERROR'; 32952 'DATA/PARAMETER MISMATCH'; 32963 'MAX CONNECTIONS EXCEEDED'; 32964 'FIREWALL'; 65535 'STATE: DISCONNECT'; 32966 'PARTNER UNAVAILABLE'; -1 'NO STATE'; 32965 'CONNECTION REFUSED'

text list "Disconnect Code Descriptions Short": 0 'DISCONNECTION SUCCESSFUL'; 28672 'NO JOB'; 28673 'JOB STARTED'; 28674 'REQUEST DURING EXECUTION'; 32902 'ID INVALID: OUT OF RANGE'; 32931 'CONNECTION ALREADY TERMINATED'; 32964 'REQUEST DURING PARAM ASSIGNMENT'; 65535 'STATE: CONNECT'; -1 'NO STATE'

text list "Text List Select": 0 ''; 1 ''; 2 ''; 3 ''

ScreenModuleEditorView "Connection_Status_Element" 392x110
   TextField "operation_label" at 0,0 size 110x110; Text 'S'
      Visibility <- "interface.operation_label_visible"
      Appearance <- "interface.operation_label_animate"
   TextField "done_status_indicator" at 110,0 size 94x27; Text 'DONE'
      Visibility <- "interface.done_status_indicator_visible"
      Appearance <- "interface.done_status_indicator_animate"
   TextField "busy_status_indicator" at 204,0 size 94x27; Text 'BUSY'
      Visibility <- "interface.busy_status_indicator_visible"
      Appearance <- "interface.busy_status_indicator_animate"
   TextField "error_status_indicator" at 298,0 size 94x27; Text 'ERROR'
      Visibility <- "interface.error_status_indicator_visible"
      Appearance <- "interface.error_status_indicator_animate"
   TextField "status_code_label" at 110,27 size 82x28; Text 'CODE:'
      Visibility <- "interface.status_code_label_visible"
      Appearance <- "interface.status_code_label_animate"
   IOField "status_code" at 192,27 size 200x28; FormatPattern ??????
      Appearance <- "interface.status_code_value_animate"
      Visibility <- "interface.status_code_value_visible"
      ProcessValue <- "interface.status_code_value"
   SymbolicIOField "status_description" at 110,55 size 282x55; TextOn '1'; TextOff '0'; TextList "Text List Select"
      Appearance <- "interface.status_code_description_animate"
      ProcessValue <- "operation_list_selector"
      Visibility <- "interface.status_code_description_visible"
   Button "operation_left" at 0,0 size 110x110; TextOff 'Text'
      on Press: function_b14e0dd5("interface.operation_button_actuate", 0)
      Visibility <- "interface.operation_button_visible"
      ObjectEnable <- "interface.operation_button_enable"
   Button "show_status" at 110,0 size 282x110; TextOff 'Text'
      on Press: function_b14e0dd5("interface.show_status_code_description_button_actuate", 0)
      Visibility <- "interface.show_status_code_description_button_visible"
      ObjectEnable <- "interface.show_status_code_description_button_enable"
*)

(* ===== HMI "HMI_RT_1" =====
system functions are stored by id; their names below are inferred from use

